(* Logix 5000 project; controller PLC_MCC1300_75F1 vendor 1 type 14 code 166 rev 32.11; software revision 32.04; part 33 of 83 *)
(* tags used below, declared in another part *)
   BENCH_MASTERUP : ALIAS FOR I[73].6;
   I : INT[128];   // Local Input Updates Input Slot 2
   KD_N_MOVIN : ALIAS FOR N14[256].0;
   KD_N_MOVOUT : ALIAS FOR N14[257].0;
   KD_S_MOVIN : ALIAS FOR N14[256].1;
   KD_S_MOVOUT : ALIAS FOR N14[257].1;
   KK_N_MOVDN : ALIAS FOR N14[253].0;
   KK_N_MOVIN : ALIAS FOR N14[254].0;
   KK_N_MOVOUT : ALIAS FOR N14[255].0;
   KK_N_MOVUP : ALIAS FOR N14[252].0;
   KK_S_MOVDN : ALIAS FOR N14[253].1;
   KK_S_MOVIN : ALIAS FOR N14[254].1;
   KK_S_MOVOUT : ALIAS FOR N14[255].1;
   KK_S_MOVUP : ALIAS FOR N14[252].1;
   KNRL_K_NTH_ADJ : ALIAS FOR O[19].0;
   KNRL_K_STH_ADJ : ALIAS FOR O[19].1;
   KNRL_N_AUTO : ALIAS FOR N14[250].0;
   KNRL_N_MANL : ALIAS FOR N14[251].0;
   KNRL_S_AUTO : ALIAS FOR N14[250].1;
   KNRL_S_MANL : ALIAS FOR N14[251].1;
   KNRL_T_NTH_ADJ : ALIAS FOR O[22].0;
   KNRL_T_STH_ADJ : ALIAS FOR O[22].1;
   N14 : DINT[500];
   O : INT[128];
   TD1_N_MOVIN : ALIAS FOR N14[256].2;
   TD1_N_MOVOUT : ALIAS FOR N14[257].2;
   TD1_S_MOVIN : ALIAS FOR N14[256].3;
   TD1_S_MOVOUT : ALIAS FOR N14[257].3;
   TD2_N_MOVIN : ALIAS FOR N14[256].4;
   TD2_N_MOVOUT : ALIAS FOR N14[257].4;
   TD2_S_MOVIN : ALIAS FOR N14[256].5;
   TD2_S_MOVOUT : ALIAS FOR N14[257].5;
   TD3_N_MOVIN : ALIAS FOR N14[256].6;
   TD3_N_MOVOUT : ALIAS FOR N14[257].6;
   TD3_S_MOVIN : ALIAS FOR N14[256].7;
   TD3_S_MOVOUT : ALIAS FOR N14[257].7;
   TD4_N_MOVIN : ALIAS FOR N14[256].8;
   TD4_N_MOVOUT : ALIAS FOR N14[257].8;
   TD4_S_MOVIN : ALIAS FOR N14[256].9;
   TD4_S_MOVOUT : ALIAS FOR N14[257].9;
   TD5_N_MOVIN : ALIAS FOR N14[256].10;
   TD5_N_MOVOUT : ALIAS FOR N14[257].10;
   TD5_S_MOVIN : ALIAS FOR N14[256].11;
   TD5_S_MOVOUT : ALIAS FOR N14[257].11;
   TDN_FLT : ALIAS FOR I[18].1;
   TDN_FWD : ALIAS FOR O[20].1;
   TDN_REV : ALIAS FOR O[20].5;
   TDN_SS1 : ALIAS FOR O[20].13;
   TDN_SS2 : ALIAS FOR O[20].9;
   TDS_FLT : ALIAS FOR I[18].2;
   TDS_FWD : ALIAS FOR O[20].2;
   TDS_REV : ALIAS FOR O[20].6;
   TDS_SS1 : ALIAS FOR O[20].14;
   TDS_SS2 : ALIAS FOR O[20].10;
   TK1_N_MOVDN : ALIAS FOR N14[253].2;
   TK1_N_MOVIN : ALIAS FOR N14[254].2;
   TK1_N_MOVOUT : ALIAS FOR N14[255].2;
   TK1_N_MOVUP : ALIAS FOR N14[252].2;
   TK1_S_MOVDN : ALIAS FOR N14[253].3;
   TK1_S_MOVIN : ALIAS FOR N14[254].3;
   TK1_S_MOVOUT : ALIAS FOR N14[255].3;
   TK1_S_MOVUP : ALIAS FOR N14[252].3;
   TK2_N_MOVDN : ALIAS FOR N14[253].4;
   TK2_N_MOVIN : ALIAS FOR N14[254].4;
   TK2_N_MOVOUT : ALIAS FOR N14[255].4;
   TK2_N_MOVUP : ALIAS FOR N14[252].4;
   TK2_S_MOVDN : ALIAS FOR N14[253].5;
   TK2_S_MOVIN : ALIAS FOR N14[254].5;
   TK2_S_MOVOUT : ALIAS FOR N14[255].5;
   TK2_S_MOVUP : ALIAS FOR N14[252].5;
   TK3_N_MOVDN : ALIAS FOR N14[253].6;
   TK3_N_MOVIN : ALIAS FOR N14[254].6;
   TK3_N_MOVOUT : ALIAS FOR N14[255].6;
   TK3_N_MOVUP : ALIAS FOR N14[252].6;
   TK3_S_MOVDN : ALIAS FOR N14[253].7;
   TK3_S_MOVIN : ALIAS FOR N14[254].7;
   TK3_S_MOVOUT : ALIAS FOR N14[255].7;
   TK3_S_MOVUP : ALIAS FOR N14[252].7;
   TK4_N_MOVDN : ALIAS FOR N14[253].8;
   TK4_N_MOVIN : ALIAS FOR N14[254].8;
   TK4_N_MOVOUT : ALIAS FOR N14[255].8;
   TK4_N_MOVUP : ALIAS FOR N14[252].8;
   TK4_S_MOVDN : ALIAS FOR N14[253].9;
   TK4_S_MOVIN : ALIAS FOR N14[254].9;
   TK4_S_MOVOUT : ALIAS FOR N14[255].9;
   TK4_S_MOVUP : ALIAS FOR N14[252].9;
   TK5_N_MOVDN : ALIAS FOR N14[253].10;
   TK5_N_MOVIN : ALIAS FOR N14[254].10;
   TK5_N_MOVOUT : ALIAS FOR N14[255].10;
   TK5_N_MOVUP : ALIAS FOR N14[252].10;
   TK5_S_MOVDN : ALIAS FOR N14[253].11;
   TK5_S_MOVIN : ALIAS FOR N14[254].11;
   TK5_S_MOVOUT : ALIAS FOR N14[255].11;
   TK5_S_MOVUP : ALIAS FOR N14[252].11;
   TK_FLT : ALIAS FOR I[18].0;
   TK_FWD : ALIAS FOR O[20].0;
   TK_REV : ALIAS FOR O[20].4;
   TK_SS1 : ALIAS FOR O[20].12;
   TK_SS2 : ALIAS FOR O[20].8;
   TZ1_K_NTH_ADJ : ALIAS FOR O[19].2;
   TZ1_K_STH_ADJ : ALIAS FOR O[19].3;
   TZ1_N_AUTO : ALIAS FOR N14[250].2;
   TZ1_N_MANL : ALIAS FOR N14[251].2;
   TZ1_S_AUTO : ALIAS FOR N14[250].3;
   TZ1_S_MANL : ALIAS FOR N14[251].3;
   TZ1_T_NTH_ADJ : ALIAS FOR O[22].2;
   TZ1_T_STH_ADJ : ALIAS FOR O[22].3;
   TZ2_K_NTH_ADJ : ALIAS FOR O[19].4;
   TZ2_K_STH_ADJ : ALIAS FOR O[19].5;
   TZ2_N_AUTO : ALIAS FOR N14[250].4;
   TZ2_N_MANL : ALIAS FOR N14[251].4;
   TZ2_S_AUTO : ALIAS FOR N14[250].5;
   TZ2_S_MANL : ALIAS FOR N14[251].5;
   TZ2_T_NTH_ADJ : ALIAS FOR O[22].4;
   TZ2_T_STH_ADJ : ALIAS FOR O[22].5;
   TZ3_K_NTH_ADJ : ALIAS FOR O[19].6;
   TZ3_K_STH_ADJ : ALIAS FOR O[19].7;
   TZ3_N_AUTO : ALIAS FOR N14[250].6;
   TZ3_N_MANL : ALIAS FOR N14[251].6;
   TZ3_S_AUTO : ALIAS FOR N14[250].7;
   TZ3_S_MANL : ALIAS FOR N14[251].7;
   TZ3_T_NTH_ADJ : ALIAS FOR O[22].6;
   TZ3_T_STH_ADJ : ALIAS FOR O[22].7;
   TZ4_K_NTH_ADJ : ALIAS FOR O[19].8;
   TZ4_K_STH_ADJ : ALIAS FOR O[19].9;
   TZ4_N_AUTO : ALIAS FOR N14[250].8;
   TZ4_N_MANL : ALIAS FOR N14[251].8;
   TZ4_S_AUTO : ALIAS FOR N14[250].9;
   TZ4_S_MANL : ALIAS FOR N14[251].9;
   TZ4_T_NTH_ADJ : ALIAS FOR O[22].8;
   TZ4_T_STH_ADJ : ALIAS FOR O[22].9;
   TZ5_K_NTH_ADJ : ALIAS FOR O[19].10;
   TZ5_K_STH_ADJ : ALIAS FOR O[19].11;
   TZ5_N_AUTO : ALIAS FOR N14[250].10;
   TZ5_N_MANL : ALIAS FOR N14[251].10;
   TZ5_S_AUTO : ALIAS FOR N14[250].11;
   TZ5_S_MANL : ALIAS FOR N14[251].11;
   TZ5_T_NTH_ADJ : ALIAS FOR O[22].10;
   TZ5_T_STH_ADJ : ALIAS FOR O[22].11;
(* MainProgram, continued *)

ROUTINE _71_LADDER   (* ladder *)
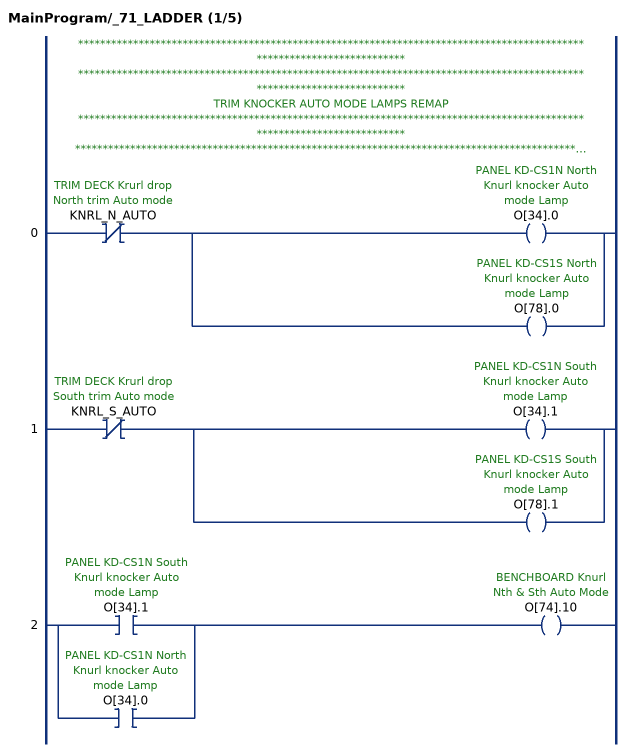
   // ***********************************************************************************************************************
   // ***********************************************************************************************************************
   //                                             TRIM KNOCKER AUTO MODE LAMPS REMAP
   // ***********************************************************************************************************************
   // ***********************************************************************************************************************
   // Knurl knocker auto mode lamps
   0: XIO(KNRL_N_AUTO)[OTE(O[34].0) ,OTE(O[78].0) ];
   1: XIO(KNRL_S_AUTO)[OTE(O[34].1) ,OTE(O[78].1) ];
   2: [XIC(O[34].1) ,XIC(O[34].0) ]OTE(O[74].10);
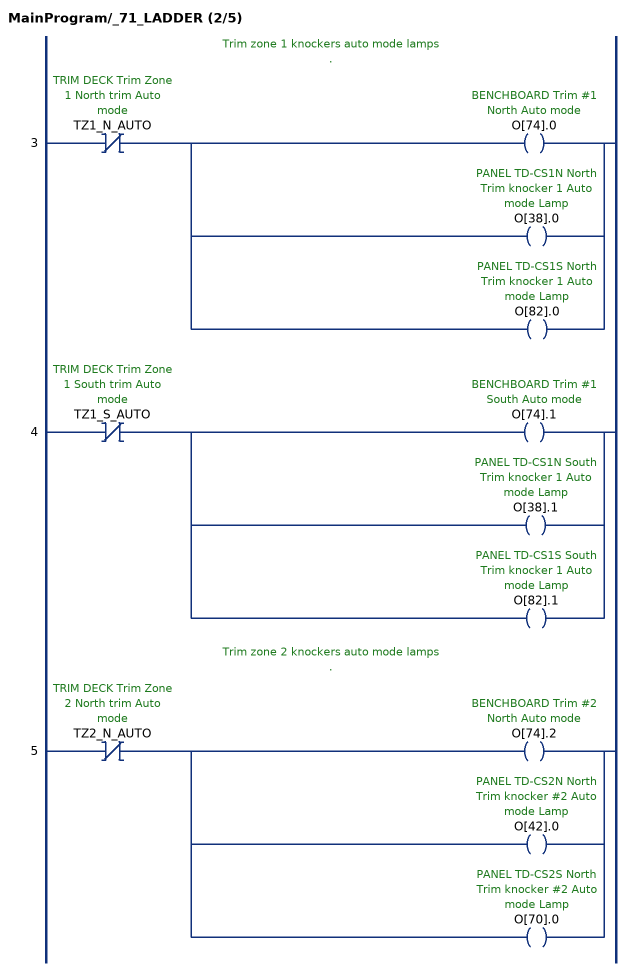
   // Trim zone 1 knockers auto mode lamps
   //                                                                                   .
   3: XIO(TZ1_N_AUTO)[OTE(O[74].0) ,OTE(O[38].0) ,OTE(O[82].0) ];
   4: XIO(TZ1_S_AUTO)[OTE(O[74].1) ,OTE(O[38].1) ,OTE(O[82].1) ];
   // Trim zone 2 knockers auto mode lamps
   //                                                                                   .
   5: XIO(TZ2_N_AUTO)[OTE(O[74].2) ,OTE(O[42].0) ,OTE(O[70].0) ];
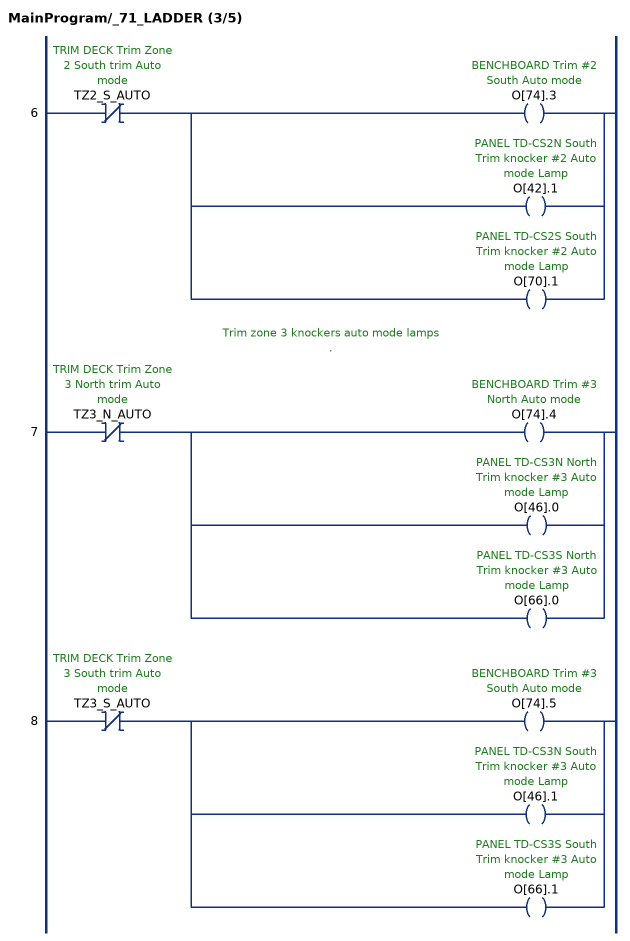
   6: XIO(TZ2_S_AUTO)[OTE(O[74].3) ,OTE(O[42].1) ,OTE(O[70].1) ];
   // Trim zone 3 knockers auto mode lamps
   //                                                                                   .
   7: XIO(TZ3_N_AUTO)[OTE(O[74].4) ,OTE(O[46].0) ,OTE(O[66].0) ];
   8: XIO(TZ3_S_AUTO)[OTE(O[74].5) ,OTE(O[46].1) ,OTE(O[66].1) ];
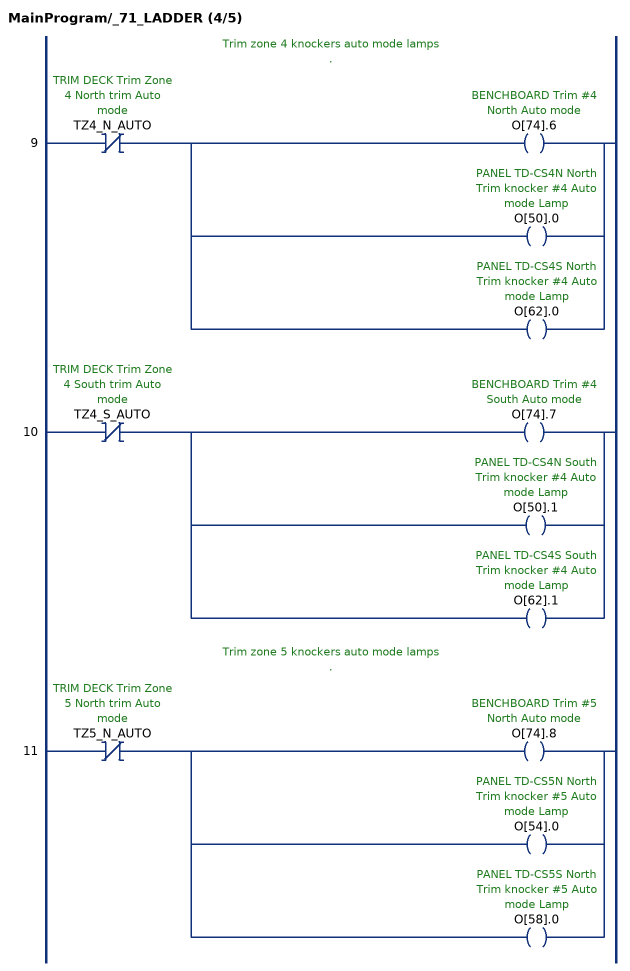
   // Trim zone 4 knockers auto mode lamps
   //                                                                                   .
   9: XIO(TZ4_N_AUTO)[OTE(O[74].6) ,OTE(O[50].0) ,OTE(O[62].0) ];
   10: XIO(TZ4_S_AUTO)[OTE(O[74].7) ,OTE(O[50].1) ,OTE(O[62].1) ];
   // Trim zone 5 knockers auto mode lamps
   //                                                                                   .
   11: XIO(TZ5_N_AUTO)[OTE(O[74].8) ,OTE(O[54].0) ,OTE(O[58].0) ];
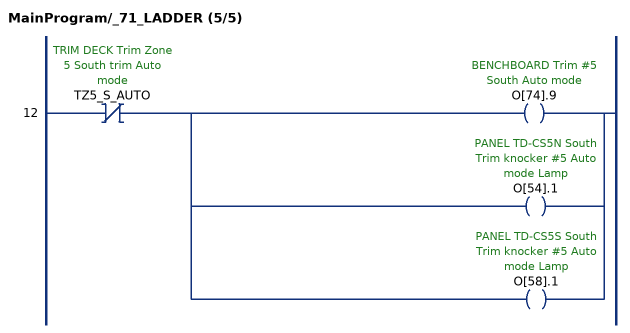
   12: XIO(TZ5_S_AUTO)[OTE(O[74].9) ,OTE(O[54].1) ,OTE(O[58].1) ];
END_ROUTINE

ROUTINE _72_LADDER   (* ladder *)
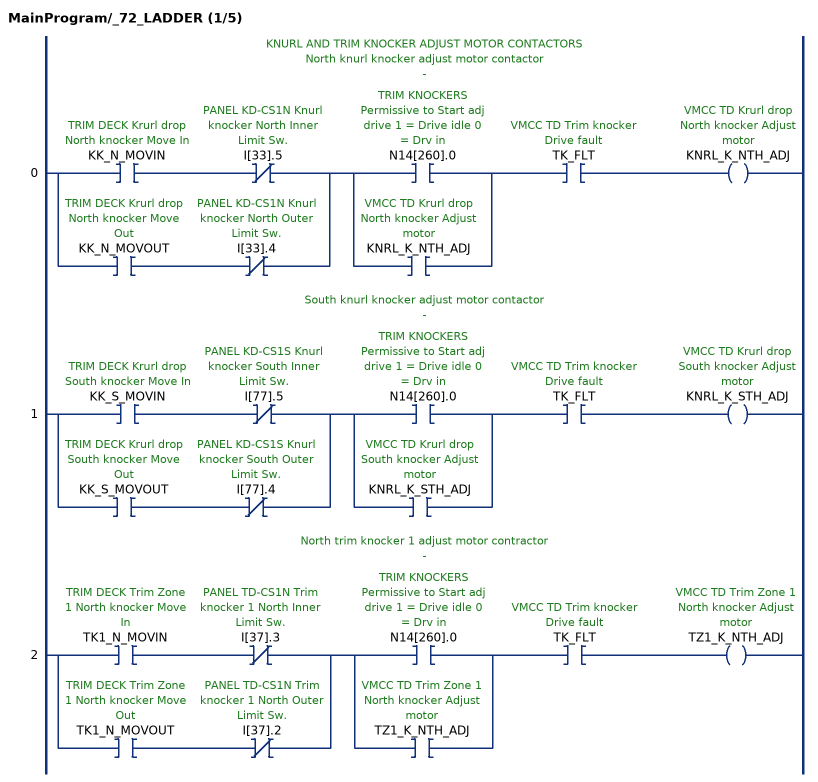
   // KNURL AND TRIM KNOCKER ADJUST MOTOR CONTACTORS
   // North knurl knocker adjust motor contactor
   //                                               -
   0: [XIC(KK_N_MOVIN) XIO(I[33].5) ,XIC(KK_N_MOVOUT) XIO(I[33].4) ][XIC(N14[260].0) ,XIC(KNRL_K_NTH_ADJ) ]XIC(TK_FLT)OTE(KNRL_K_NTH_ADJ);
   // South knurl knocker adjust motor contactor
   //                                               -
   1: [XIC(KK_S_MOVIN) XIO(I[77].5) ,XIC(KK_S_MOVOUT) XIO(I[77].4) ][XIC(N14[260].0) ,XIC(KNRL_K_STH_ADJ) ]XIC(TK_FLT)OTE(KNRL_K_STH_ADJ);
   // North trim knocker 1 adjust motor contractor
   //                                                            -
   2: [XIC(TK1_N_MOVIN) XIO(I[37].3) ,XIC(TK1_N_MOVOUT) XIO(I[37].2) ][XIC(N14[260].0) ,XIC(TZ1_K_NTH_ADJ) ]XIC(TK_FLT)OTE(TZ1_K_NTH_ADJ);
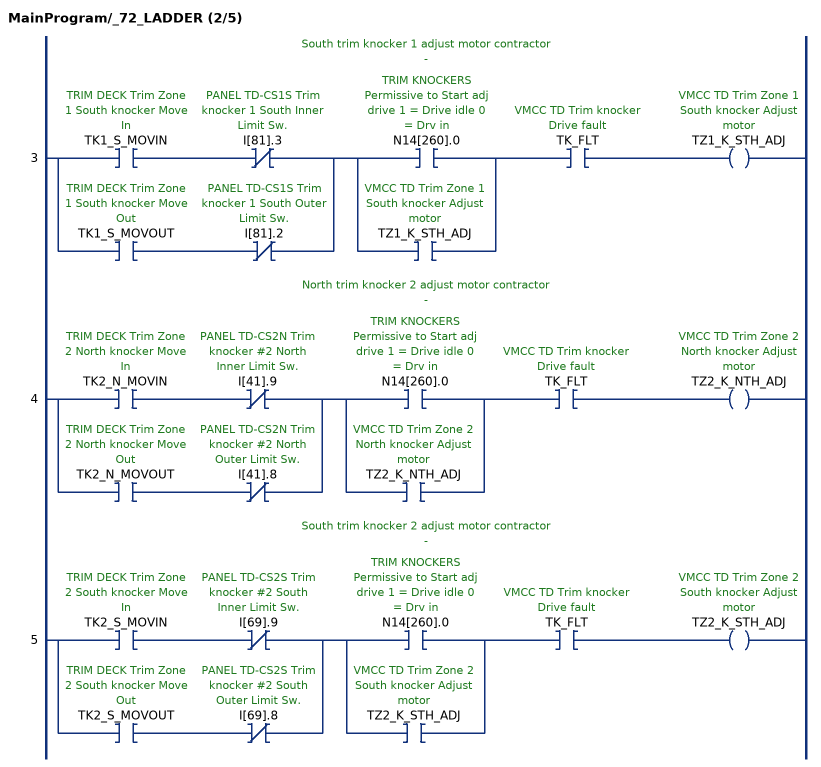
   // South trim knocker 1 adjust motor contractor
   //                                                                           -
   3: [XIC(TK1_S_MOVIN) XIO(I[81].3) ,XIC(TK1_S_MOVOUT) XIO(I[81].2) ][XIC(N14[260].0) ,XIC(TZ1_K_STH_ADJ) ]XIC(TK_FLT)OTE(TZ1_K_STH_ADJ);
   // North trim knocker 2 adjust motor contractor
   //                                                                   -
   4: [XIC(TK2_N_MOVIN) XIO(I[41].9) ,XIC(TK2_N_MOVOUT) XIO(I[41].8) ][XIC(N14[260].0) ,XIC(TZ2_K_NTH_ADJ) ]XIC(TK_FLT)OTE(TZ2_K_NTH_ADJ);
   // South trim knocker 2 adjust motor contractor
   //                                                                       -
   5: [XIC(TK2_S_MOVIN) XIO(I[69].9) ,XIC(TK2_S_MOVOUT) XIO(I[69].8) ][XIC(N14[260].0) ,XIC(TZ2_K_STH_ADJ) ]XIC(TK_FLT)OTE(TZ2_K_STH_ADJ);
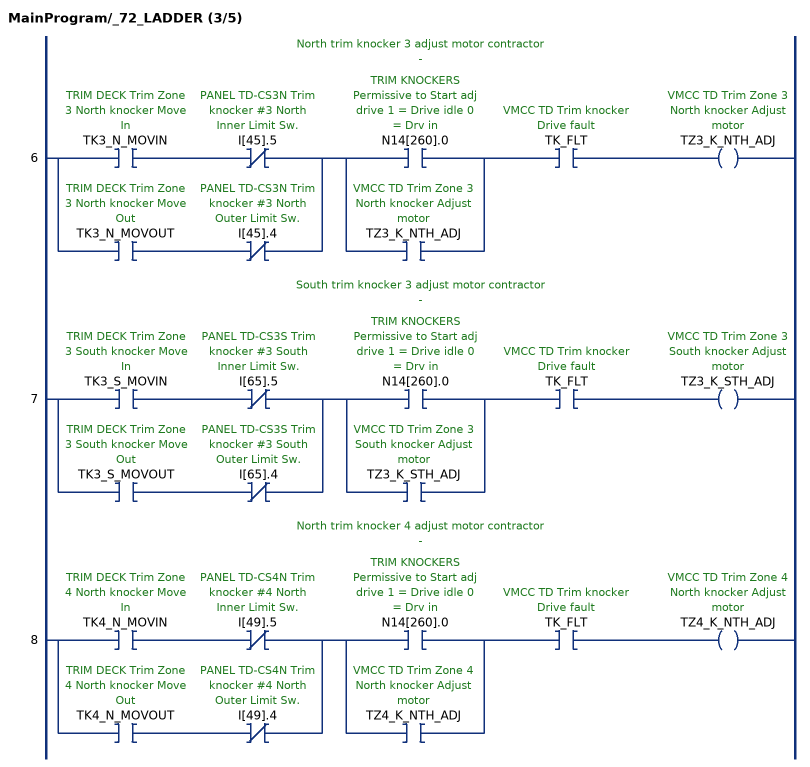
   // North trim knocker 3 adjust motor contractor
   //                                                                       -
   6: [XIC(TK3_N_MOVIN) XIO(I[45].5) ,XIC(TK3_N_MOVOUT) XIO(I[45].4) ][XIC(N14[260].0) ,XIC(TZ3_K_NTH_ADJ) ]XIC(TK_FLT)OTE(TZ3_K_NTH_ADJ);
   // South trim knocker 3 adjust motor contractor
   //                                                                       -
   7: [XIC(TK3_S_MOVIN) XIO(I[65].5) ,XIC(TK3_S_MOVOUT) XIO(I[65].4) ][XIC(N14[260].0) ,XIC(TZ3_K_STH_ADJ) ]XIC(TK_FLT)OTE(TZ3_K_STH_ADJ);
   // North trim knocker 4 adjust motor contractor
   //                                                                       -
   8: [XIC(TK4_N_MOVIN) XIO(I[49].5) ,XIC(TK4_N_MOVOUT) XIO(I[49].4) ][XIC(N14[260].0) ,XIC(TZ4_K_NTH_ADJ) ]XIC(TK_FLT)OTE(TZ4_K_NTH_ADJ);
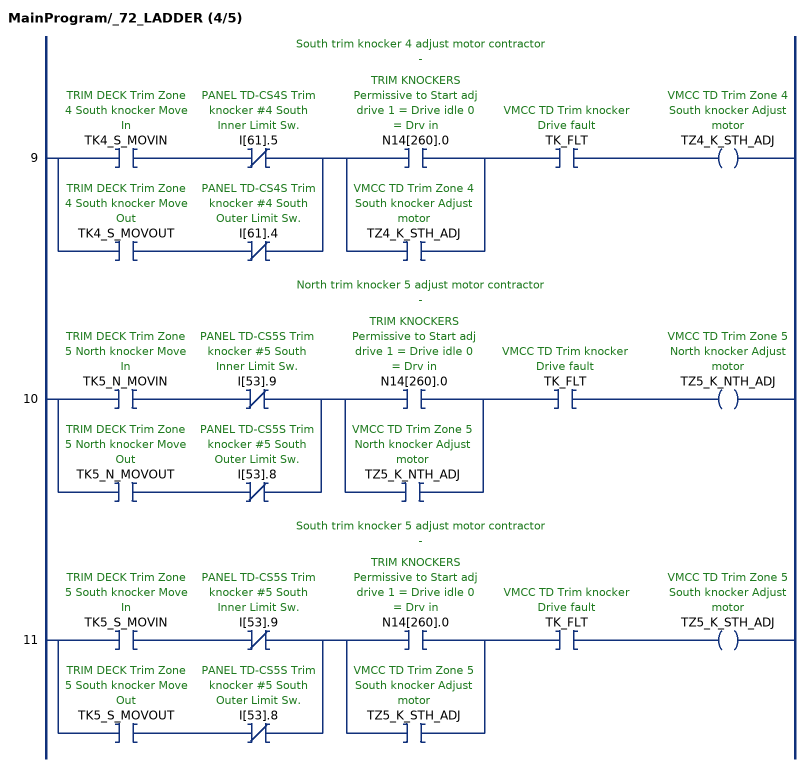
   // South trim knocker 4 adjust motor contractor
   //                                                                       -
   9: [XIC(TK4_S_MOVIN) XIO(I[61].5) ,XIC(TK4_S_MOVOUT) XIO(I[61].4) ][XIC(N14[260].0) ,XIC(TZ4_K_STH_ADJ) ]XIC(TK_FLT)OTE(TZ4_K_STH_ADJ);
   // North trim knocker 5 adjust motor contractor
   //                                                                       -
   10: [XIC(TK5_N_MOVIN) XIO(I[53].9) ,XIC(TK5_N_MOVOUT) XIO(I[53].8) ][XIC(N14[260].0) ,XIC(TZ5_K_NTH_ADJ) ]XIC(TK_FLT)OTE(TZ5_K_NTH_ADJ);
   // South trim knocker 5 adjust motor contractor
   //                                                                       -
   11: [XIC(TK5_S_MOVIN) XIO(I[53].9) ,XIC(TK5_S_MOVOUT) XIO(I[53].8) ][XIC(N14[260].0) ,XIC(TZ5_K_STH_ADJ) ]XIC(TK_FLT)OTE(TZ5_K_STH_ADJ);
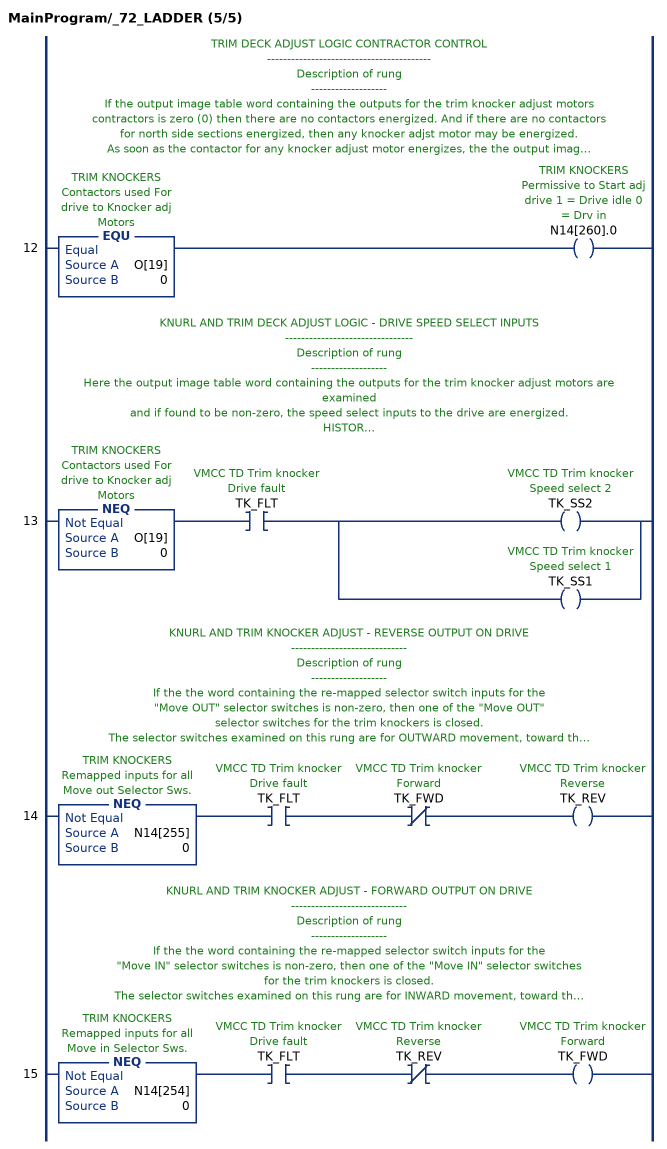
   // TRIM DECK ADJUST LOGIC CONTRACTOR CONTROL
   // -----------------------------------------
   // Description of rung
   // -------------------
   // If the output image table word containing the outputs for the trim knocker adjust motors
   // contractors is zero (0) then there are no contactors energized. And if there are no contactors
   // for north side sections energized, then any knocker adjst motor may be energized.
   // As soon as the contactor for any knocker adjust motor energizes, the the output image
   // table word containing the outputs for the trim knocker adjust motors will become non-zero.
   // HISTORY
   // =======
   // DATE        DESCRIPTION                                                       PROGRAMMER
   // ====        ===========                                                       ==========
   // 2/29/96     Entered rung as designed                                          WAS
   // 3/1/96      Entered comment                                                   WAS
   12: EQU(O[19],0)OTE(N14[260].0);
   // KNURL AND TRIM DECK ADJUST LOGIC - DRIVE SPEED SELECT INPUTS
   // --------------------------------
   // Description of rung
   // -------------------
   // Here the output image table word containing the outputs for the trim knocker adjust motors are examined
   // and if found to be non-zero, the speed select inputs to the drive are energized.
   // HISTORY
   // =======
   // DATE        DESCRIPTION                                                       PROGRAMMER
   // ====        ===========                                                       ==========
   // 2/29/96     Entered rung as designed                                          WAS
   // 3/1/96      Entered comment                                                   WAS
   13: NEQ(O[19],0)XIC(TK_FLT)[OTE(TK_SS2) ,OTE(TK_SS1) ];
   // KNURL AND TRIM KNOCKER ADJUST - REVERSE OUTPUT ON DRIVE
   // -----------------------------
   // Description of rung
   // -------------------
   // If the the word containing the re-mapped selector switch inputs for the
   // "Move OUT" selector switches is non-zero, then one of the "Move OUT"
   // selector switches for the trim knockers is closed.
   // The selector switches examined on this rung are for OUTWARD movement, toward the
   // center of the conveyors. Any movement in this direction is accomplished by operating the
   // adjust motor in the REVERSE direction. Hence, if any of the out selector switches is made, then
   // the REVERSE drive input should be energized.
   // HISTORY
   // =======
   // DATE        DESCRIPTION                                                       PROGRAMMER
   // ====        ===========                                                       ==========
   // 2/29/96     Entered rung as designed                                          WAS
   // 3/1/96      Entered comment                                                   WAS
   14: NEQ(N14[255],0)XIC(TK_FLT)XIO(TK_FWD)OTE(TK_REV);
   // KNURL AND TRIM KNOCKER ADJUST - FORWARD OUTPUT ON DRIVE
   // -----------------------------
   // Description of rung
   // -------------------
   // If the the word containing the re-mapped selector switch inputs for the
   // "Move IN" selector switches is non-zero, then one of the "Move IN" selector switches
   // for the trim knockers is closed.
   // The selector switches examined on this rung are for INWARD movement, toward the
   // center of the conveyors. Any movement in this direction is accomplished by operating the
   // adjust motor in the forward direction. Hence, if any of the out selector switches is made, then
   // the forward drive input should be energized.
   // HISTORY
   // =======
   // DATE        DESCRIPTION                                                       PROGRAMMER
   // ====        ===========                                                       ==========
   // 2/29/96     Entered rung as designed                                          WAS
   // 3/1/96      Entered comment                                                   WAS
   15: NEQ(N14[254],0)XIC(TK_FLT)XIO(TK_REV)OTE(TK_FWD);
END_ROUTINE

ROUTINE _73_LADDER   (* ladder *)
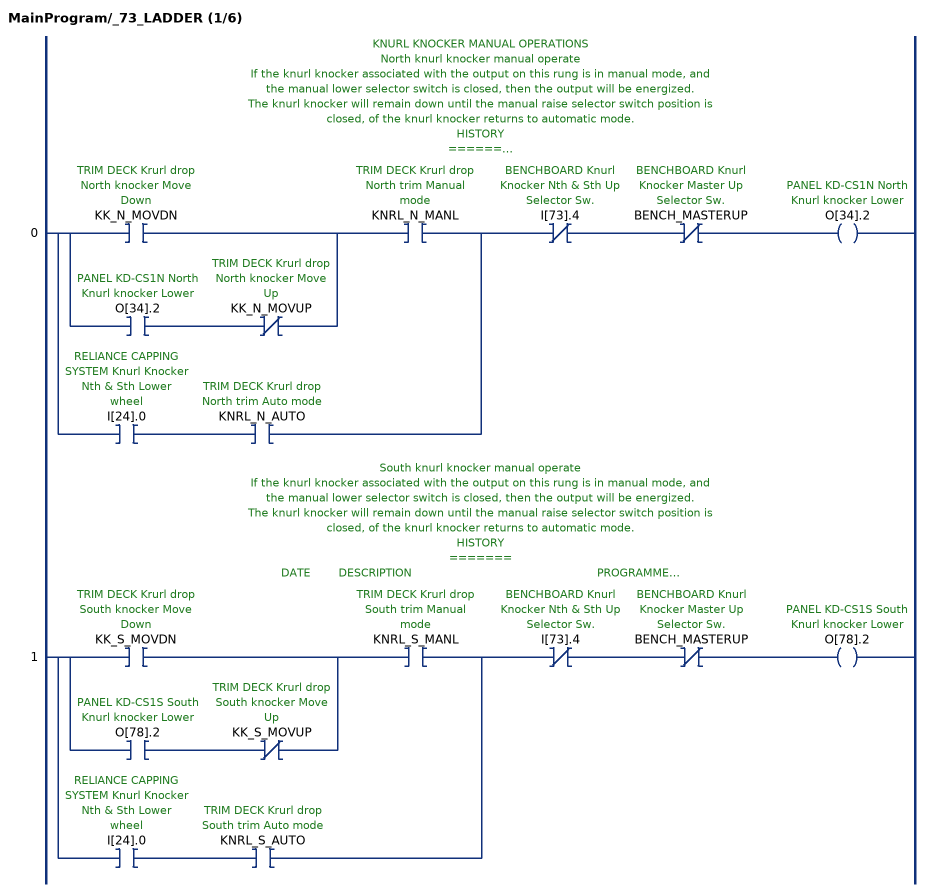
   // KNURL KNOCKER MANUAL OPERATIONS
   // North knurl knocker manual operate
   // If the knurl knocker associated with the output on this rung is in manual mode, and
   // the manual lower selector switch is closed, then the output will be energized.
   // The knurl knocker will remain down until the manual raise selector switch position is
   // closed, of the knurl knocker returns to automatic mode.
   // HISTORY
   // =======
   // DATE        DESCRIPTION                                                     PROGRAMMER
   // ====        ===========                                                     ==========
   // 2/29/96     Entered rung as designed                                        WAS
   // 3/1/96      Added these comments                                            WAS
   0: [[XIC(KK_N_MOVDN) ,XIC(O[34].2) XIO(KK_N_MOVUP) ] XIC(KNRL_N_MANL) ,XIC(I[24].0) XIC(KNRL_N_AUTO) ]XIO(I[73].4)XIO(BENCH_MASTERUP)OTE(O[34].2);
   // South knurl knocker manual operate
   // If the knurl knocker associated with the output on this rung is in manual mode, and
   // the manual lower selector switch is closed, then the output will be energized.
   // The knurl knocker will remain down until the manual raise selector switch position is
   // closed, of the knurl knocker returns to automatic mode.
   // HISTORY
   // =======
   // DATE        DESCRIPTION                                                     PROGRAMMER
   // ====        ===========                                                     ==========
   // 2/29/96     Entered rung as designed                                        WAS
   // 3/1/96      Added these comments                                            WAS
   1: [[XIC(KK_S_MOVDN) ,XIC(O[78].2) XIO(KK_S_MOVUP) ] XIC(KNRL_S_MANL) ,XIC(I[24].0) XIC(KNRL_S_AUTO) ]XIO(I[73].4)XIO(BENCH_MASTERUP)OTE(O[78].2);
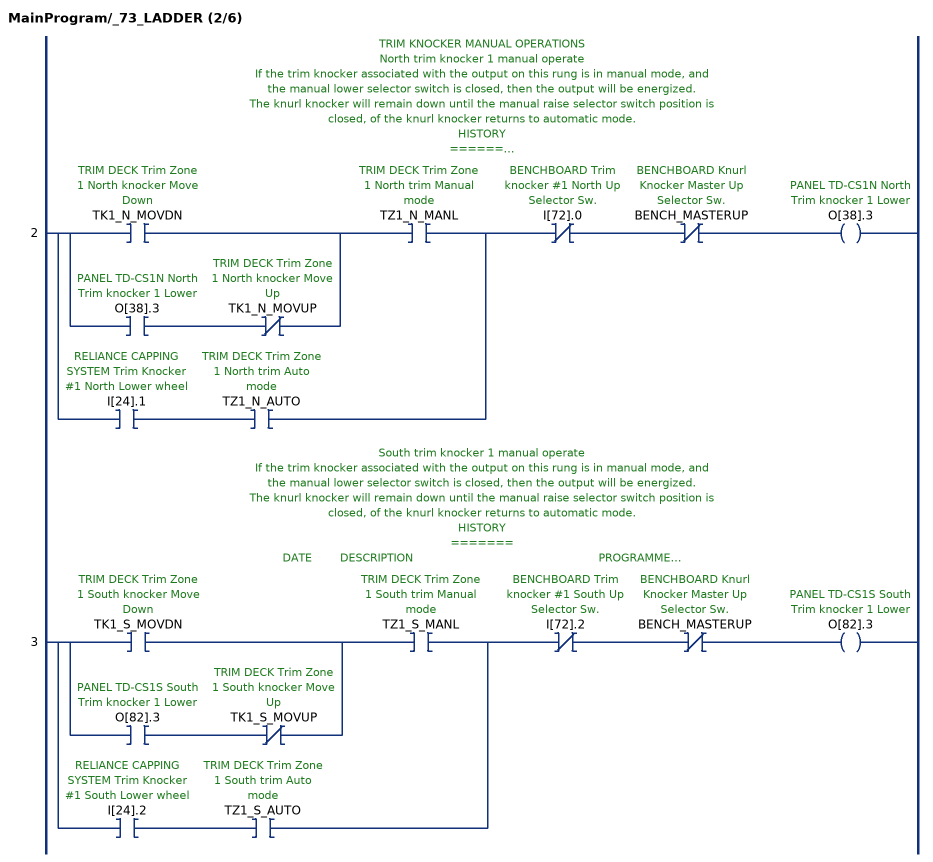
   // TRIM KNOCKER MANUAL OPERATIONS
   // North trim knocker 1 manual operate
   // If the trim knocker associated with the output on this rung is in manual mode, and
   // the manual lower selector switch is closed, then the output will be energized.
   // The knurl knocker will remain down until the manual raise selector switch position is
   // closed, of the knurl knocker returns to automatic mode.
   // HISTORY
   // =======
   // DATE        DESCRIPTION                                                     PROGRAMMER
   // ====        ===========                                                     ==========
   // 2/29/96     Entered rung as designed                                        WAS
   // 3/1/96      Added these comments                                            WAS
   2: [[XIC(TK1_N_MOVDN) ,XIC(O[38].3) XIO(TK1_N_MOVUP) ] XIC(TZ1_N_MANL) ,XIC(I[24].1) XIC(TZ1_N_AUTO) ]XIO(I[72].0)XIO(BENCH_MASTERUP)OTE(O[38].3);
   // South trim knocker 1 manual operate
   // If the trim knocker associated with the output on this rung is in manual mode, and
   // the manual lower selector switch is closed, then the output will be energized.
   // The knurl knocker will remain down until the manual raise selector switch position is
   // closed, of the knurl knocker returns to automatic mode.
   // HISTORY
   // =======
   // DATE        DESCRIPTION                                                     PROGRAMMER
   // ====        ===========                                                     ==========
   // 2/29/96     Entered rung as designed                                        WAS
   // 3/1/96      Added these comments                                            WAS
   3: [[XIC(TK1_S_MOVDN) ,XIC(O[82].3) XIO(TK1_S_MOVUP) ] XIC(TZ1_S_MANL) ,XIC(I[24].2) XIC(TZ1_S_AUTO) ]XIO(I[72].2)XIO(BENCH_MASTERUP)OTE(O[82].3);